(* Logix 5000 project; controller Digital_Interlock_PLC vendor 1 type 14 code 196 rev 37.11; software revision 37.00 *) (continued)
ADD_ON_INSTRUCTION AOI_Sys_Module   (* revision 1.0, vendor Jeremy Medders, ExecutePrescan *)
// Provides detailed module diagnostics and inhibit ability.
VAR_IN_OUT
   Ref_Module : MODULE; {required}   // Name of the module in the I/O tree.
END_VAR
VAR_INPUT
   Inp_Inhibit : BOOL; {access Read Only, visible}   // Command to inhibit the module.
   Inp_Uninhibit : BOOL; {access Read Only, visible}   // Command to uninhibit the module.
END_VAR
VAR_OUTPUT
   Val_EntryStatus : DINT; {access Read Only, visible}   // Specifies the current state of the specified map entry.
   Val_FaultCode : DINT; {access Read Only, visible}   // A number that identifies a module fault, if one occurs.
   Val_FaultInfo : DINT; {access Read Only, visible}   // Provides specific information about the Module object fault code.
   Val_Instance : DINT; {access Read Only, visible}   // Provides the instance number of this module object.
   Val_Mode : DINT; {access Read Only, visible}   // Specifies the current mode of the Module object.
   Sts_Standby : ALIAS FOR Status.0; {access Read Only, visible}   // The controller is powering up.
   Sts_Faulted : ALIAS FOR Status.1; {access Read Only, visible}   // Indicates whether any of the Module object’s connections to the associated module have failed.
   Sts_Validating : ALIAS FOR Status.2; {access Read Only, visible}   // The Module object is verifying Module object integrity prior to establishing connections to the module.
   Sts_Connecting : ALIAS FOR Status.3; {access Read Only, visible}   // The Module object is initiating connections to the module.
   Sts_Connected : ALIAS FOR Status.4; {access Read Only, visible}   // All connections to the module are established and data is transferring.
   Sts_ShuttingDown : ALIAS FOR Status.5; {access Read Only, visible}   // The Module object is in the process of shutting down all connections to the module.
   Sts_Inhibited : ALIAS FOR Status.6; {access Read Only, visible}   // The Module object is inhibited (the inhibit bit in the Mode attribute is set).
   Sts_Waiting : ALIAS FOR Status.7; {access Read Only, visible}   // The parent object upon which this Module object depends is not running.
   Sts_FirmwareUpdating : ALIAS FOR Status.9; {access Read Only, visible}   // Firmware supervisor is attempting to flash the module.
   Sts_Configuring : ALIAS FOR Status.10; {access Read Only, visible}   // Controller is downloading configuration to the module.
   Sts_Disconnected : ALIAS FOR Status.11; {access Read Only, visible}
END_VAR
VAR
   ModeSet : DINT; {access None}
   OSR : BOOL; {access None}
   ESts : DINT; {access None}
   Status : DINT; {access Read Only}
END_VAR

ROUTINE Logic   (* structured text *)
   
   /*
       AO_Sys_Module
       Purpose:
         - Read a module object's status, fault info, and mode
         - One-shot inhibit/uninhibit via Mode bit 2 (0x0004)
         - Decode EntryStatus into HMI-friendly booleans
   */
   
   // --- Snapshot current module diagnostics/state ---
   GSV(Module, Ref_Module, INSTANCE, Val_Instance);
   GSV(Module, Ref_Module, EntryStatus, Val_EntryStatus);
   GSV(Module, Ref_Module, FaultCode, Val_FaultCode);
   GSV(Module, Ref_Module, FaultInfo, Val_FaultInfo);
   GSV(Module, Ref_Module, Mode, Val_Mode);
   
   // --- Rising-edge one-shots for inhibit control (bit 2 of Mode) ---
   // Inhibit: set bit 2
   if (Inp_Inhibit & NOT OSR) then
   	ModeSet := Val_Mode OR 16#0004;
   	SSV(Module, Ref_Module, Mode, ModeSet);
   
   // Uninhibit: clear bit 2
   elsif (Inp_Uninhibit & NOT OSR) then
   	ModeSet := Val_Mode AND 16#FFFB;
   	SSV(Module, Ref_Module, Mode, ModeSet);
   end_if;
   
   // One-shot memory: true for one scan when either command goes high
   OSR := Inp_Inhibit OR Inp_Uninhibit;
   
   /*
   	Entry Status Map
   	• 0x0000: Standby
   	• 0x1000: Faulted
   	• 0x2000: Validating
   	• 0x3000: Connecting
   	• 0x4000: Running
   	• 0x5000: Shutting Down
   	• 0x6000: Inhibited
   	• 0x7000: Waiting
   	• 0x9000: Firmware Updating
   	• 0xA000: Configuring
   */
   ESts := Val_EntryStatus & 16#F000;
   
   // State booleans for HMI/logic
   Sts_Standby := (ESts = 16#0000);
   Sts_Faulted := (ESts = 16#1000);
   Sts_Validating := (ESts = 16#2000);
   Sts_Connecting := (ESts = 16#3000);
   Sts_Connected := (ESts = 16#4000);
   Sts_ShuttingDown := (ESts = 16#5000);
   Sts_Inhibited := (ESts = 16#6000);
   Sts_Waiting := (ESts = 16#7000);
   Sts_FirmwareUpdating := (ESts = 16#9000);
   Sts_Configuring := (ESts = 16#A000);
   Sts_Disconnected := NOT (Sts_Inhibited OR Sts_Connected);
   
END_ROUTINE

ROUTINE Prescan   (* structured text *)
   
   /*
   	AO_Sys_Module
   */
   
   Inp_Inhibit := 0;
   Inp_Uninhibit := 0;
   
   Status := 0;
   
   Val_Instance := 0;
   Val_EntryStatus := 0;
   Val_FaultCode := 0;
   Val_FaultInfo := 0;
   Val_Mode := 0;
   
END_ROUTINE
END_ADD_ON_INSTRUCTION

VAR_GLOBAL   (* controller tags *)
   _DEBUG : BOOL;
   CommsStatus : DINT;
        .3   // LIC comms ok
        .0   // Prefeeder comms ok
        .1   // Stacker comms ok
        .2   // Press comms ok
   CommsStatus_Prefeeder : DINT := 11;
   CommsStatus_Press : DINT;
   CommsStatus_Stacker : DINT;
   EnableLineOptimization : BOOL;
   FaultDetected : BOOL;   // Bool to execute fault routine
   FeedInterruptActive : BOOL;
   FromLIC : UDT_FromLIC;   // Data received from LIC Client
   FromPrefeeder : UDT_EIP_FromPrefeeder;
   FromPress : UDT_EIP_FromPress;
   FromStacker : UDT_EIP_FromStacker;
   HB_ScanCounter : INT := 50;
   HB_Timer1 : TIMER := (PRE := 20);
   HB_Timer2 : TIMER := (PRE := 20);
   HeartBeat : DINT;
   MachineCount : DINT;
   PF_MSG : MESSAGE;
        MessageParameters(ServiceCode := 16#004d, LocalElement := ToPrefeeder.Heartbeat, ...)
   State : UDT_StateContext;
   States : UDT_States;
   ToLIC : UDT_ToLIC;   // Data sent to LIC Client
   ToPrefeeder : UDT_EIP_ToPrefeeder := (Heartbeat := 27);
   ToPress : UDT_EIP_ToPress;
   ToStacker : UDT_EIP_ToStacker := (PrintStation[0].blnSideWaysActive := 1);
END_VAR

PROGRAM Fault_Handler_Program   (* main routine ControllerFaultHandlerRoutine, fault routine CheckSpecificFaultRoutine *)
VAR
   CPU_Scanning : BOOL;   // Identifies when the controller is in prescan.Used t to determine if the fault occurred during prescan or normal scan of the logic
   FaultCode : DINT := 20;
   FaultType : DINT := 4;
   MajorFaultRecord : UDT_FaultRecord;
        .TimeLow   // Stores the fault information in the major_fault_record tag. When you enter a tag that is based on a structure, enter the first member of the tag
   MF_ClearRequestEnable : BOOL;   // allow program to clear this class of fault
   MF_Code : DINT;
   MF_Latched : BOOL;   // Goes true when new fault captured
   MF_Msg : STRING;
   MF_T01_C01 : STR_MajorFault := 'Major Fault T01:C01 - Power-up Fault: Power lost and restored in RUN mode. The controller that is powered on is in Run mode.'; {constant}   // The controller that is powered on is in Run mode.
   MF_T01_C16 : STR_MajorFault := 'Major Fault T01:C16 - Power-up Fault: I/O Communications Configuration fault detected.. I/O communication configuration fault detected.'; {constant}   // I/O communication configuration fault detected.
   MF_T01_C60 : STR_MajorFault := 'Major Fault T01:C60 - Power-up Fault: Non-recoverable fault. The controller detected a nonrecoverable major fault. Diagnostic information can be recovered.'; {constant}   // The controller detected a nonrecoverable major fault. Diagnostic information can be recovered.
   MF_T01_C61 : STR_MajorFault := 'Major Fault T01:C61 - Power-up Fault: Non-recoverable fault with saved diagnostic information. The controller detected a nonrecoverable major fault. Diagnostic information can be recovered.'; {constant}   // The controller detected a nonrecoverable major fault. Diagnostic information can be recovered.
   MF_T03_C16 : STR_MajorFault := 'Major Fault T03:C16 - I/O Fault: I/O module connection failed on required module. A required I/O module connection failed.'; {constant}   // A required I/O module connection failed.
   MF_T03_C23 : STR_MajorFault := 'Major Fault T03:C23 - I/O Fault: At least one required connection not established before going into RUN mode. At least one required connection was not established before going to Run mode.'; {constant}   // At least one required connection was not established before going to Run mode.
   MF_T03_C32 : STR_MajorFault := 'Major Fault T03:C32 - I/O Fault: Controller failed to open an I/O connection to a fault-tolerant I/O module because its partner controller is in a Primary state. The controller failed to open an I/O c'; {constant}   // The controller failed to open an I/O connection to a fault-tolerant I/O module because its partner controller is in a Primary state.
   MF_T03_C94 : STR_MajorFault := 'Minor Fault T03:C94 - I/O Fault: Module RPI overlap detected. The current RPI update of an I/O module overlaps with its previous RPI update.'; {constant}   // The current RPI update of an I/O module overlaps with its previous RPI update.
   MF_Timestamp : DINT;   // UTC seconds/millis, optional timestamp
   MF_Type : DINT;
END_VAR

ROUTINE CheckSpecificFaultRoutine   (* ladder *)
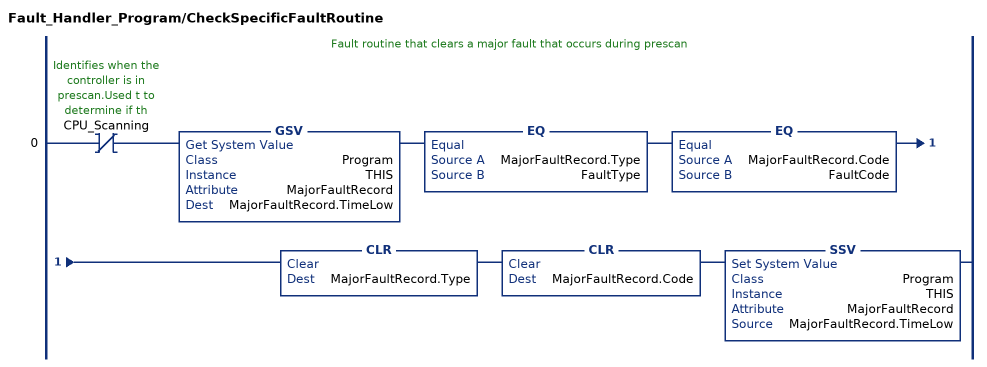
   // Fault routine that clears a major fault that occurs during prescan
   0: XIO(CPU_Scanning)GSV(Program,THIS,MajorFaultRecord,MajorFaultRecord.TimeLow)EQ(MajorFaultRecord.Type,FaultType)EQ(MajorFaultRecord.Code,FaultCode)CLR(MajorFaultRecord.Type)CLR(MajorFaultRecord.Code)SSV(Program,THIS,MajorFaultRecord,MajorFaultRecord.TimeLow);
END_ROUTINE

ROUTINE ControllerFaultHandlerRoutine   (* ladder *)
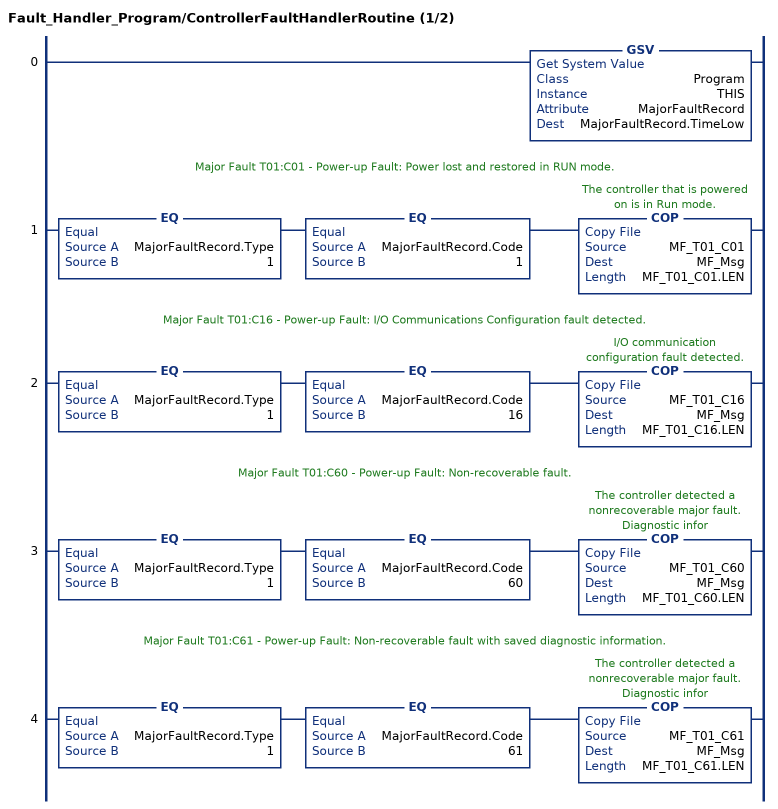
   0: GSV(Program,THIS,MajorFaultRecord,MajorFaultRecord.TimeLow);
   // Major Fault T01:C01 - Power-up Fault: Power lost and restored in RUN mode.
   1: EQ(MajorFaultRecord.Type,1)EQ(MajorFaultRecord.Code,1)COP(MF_T01_C01,MF_Msg,MF_T01_C01.LEN);
   // Major Fault T01:C16 - Power-up Fault: I/O Communications Configuration fault detected.
   2: EQ(MajorFaultRecord.Type,1)EQ(MajorFaultRecord.Code,16)COP(MF_T01_C16,MF_Msg,MF_T01_C16.LEN);
   // Major Fault T01:C60 - Power-up Fault: Non-recoverable fault.
   3: EQ(MajorFaultRecord.Type,1)EQ(MajorFaultRecord.Code,60)COP(MF_T01_C60,MF_Msg,MF_T01_C60.LEN);
   // Major Fault T01:C61 - Power-up Fault: Non-recoverable fault with saved diagnostic information.
   4: EQ(MajorFaultRecord.Type,1)EQ(MajorFaultRecord.Code,61)COP(MF_T01_C61,MF_Msg,MF_T01_C61.LEN);
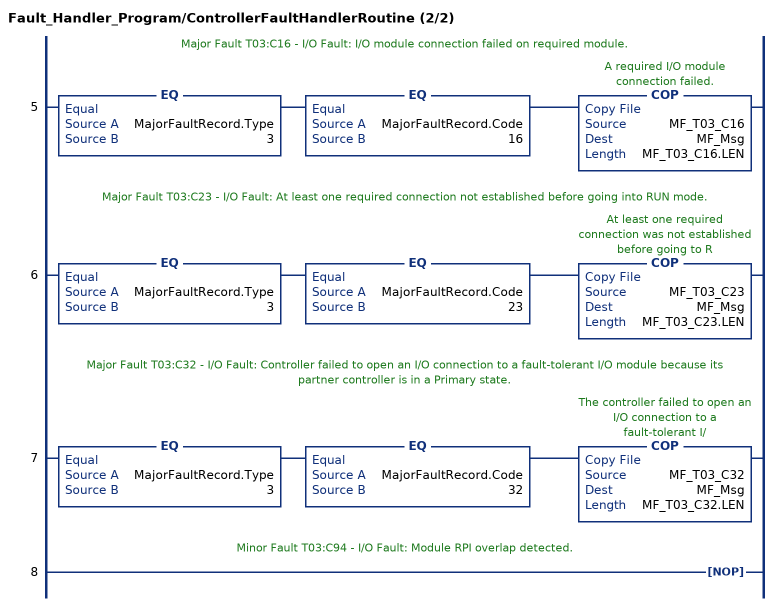
   // Major Fault T03:C16 - I/O Fault: I/O module connection failed on required module.
   5: EQ(MajorFaultRecord.Type,3)EQ(MajorFaultRecord.Code,16)COP(MF_T03_C16,MF_Msg,MF_T03_C16.LEN);
   // Major Fault T03:C23 - I/O Fault: At least one required connection not established before going into RUN mode.
   6: EQ(MajorFaultRecord.Type,3)EQ(MajorFaultRecord.Code,23)COP(MF_T03_C23,MF_Msg,MF_T03_C23.LEN);
   // Major Fault T03:C32 - I/O Fault: Controller failed to open an I/O connection to a fault-tolerant I/O module because its partner controller is in a Primary state.
   7: EQ(MajorFaultRecord.Type,3)EQ(MajorFaultRecord.Code,32)COP(MF_T03_C32,MF_Msg,MF_T03_C32.LEN);
   // Minor Fault T03:C94 - I/O Fault: Module RPI overlap detected.
   8: NOP();
END_ROUTINE
END_PROGRAM

PROGRAM MainProgram   (* main routine MainRoutine *)
VAR
   AlwaysTrue : BOOL := 1; {constant}
   AnyFault : BOOL;
   BR1_Health : UDT_DeviceHealth;
   BR2_Health : UDT_DeviceHealth;
   CmdEdge_Interrupt : BOOL;
   CmdEdge_Reconfig : BOOL;
   CmdEdge_Reset : BOOL;
   CmdEdge_Start : BOOL;
   CmdEdge_Stop : BOOL;
   CmdId_Desired : DINT;
   CmdId_Last : DINT;
   CN1_Health : UDT_DeviceHealth;
   CN2_Health : UDT_DeviceHealth;
   CommandEnum : UDT_CommandEnum;
   CommsHealthy : BOOL;   // Heartbeat Ok between peer machines
   DesiredCommand : DINT;   // From LIC Client
   EndCriteriaMet : BOOL;
   GuardsOk : BOOL;
   HeartBeatB : BOOL := 1;
   HoldClear : BOOL;
   HWReady : BOOL;   // Machines present and communicating
   MajorFaultRec : UDT_FaultRecord;
   ONS_CmdId : BOOL;
   PermissivesOk : BOOL;   // (safety, e-stops, power, guards
   PF1_Health : UDT_DeviceHealth := (DeviceConfigured := 1);
   PF2_Health : UDT_DeviceHealth;
   PL1_Health : UDT_DeviceHealth;
   PL2_Health : UDT_DeviceHealth;
   PowerOk : BOOL;
   PR1_Health : UDT_DeviceHealth;
   PR2_Health : UDT_DeviceHealth;
   SafetyChain_OK : BOOL;
   SR1_Health : UDT_DeviceHealth;
   SR2_Health : UDT_DeviceHealth;
   ST1_Health : UDT_DeviceHealth := (DeviceConfigured := 1);
   ST2_Health : UDT_DeviceHealth;
   TaskPeriod_ms : DINT := 10; {constant}   // must match periodic task ms
   TB1_Health : UDT_DeviceHealth;
   TB2_Health : UDT_DeviceHealth;
   Tmr_Hold : TIMER := (PRE := 10000);
   Tmr_Init : TIMER := (PRE := 3000);
   Tmr_Running : TIMER := (PRE := 5000);
END_VAR

ROUTINE DataRoutingRoutine   (* structured text *)
   
   /******************** 	DATA MAPPING	********************/
   
   ST1:O.Data[0] := ToStacker.Heartbeat;										// Press -> Stacker
   ST1:O.Data[1] := ToStacker.CommandedSpeed;									// Press -> Stacker
   ST1:O.Data[2] := ToStacker.PressCurrentSpeed;								// Press -> Stacker
   ST1:O.Data[3].0 := ToStacker.RollInPermissive;								// Press -> Stacker
   ST1:O.Data[3].1 := ToStacker.RunPermissive;									// Press -> Stacker
   ST1:O.Data[3].2 := ToStacker.VOSReset;										// Press -> Stacker
   ST1:O.Data[3].3 := ToStacker.VOSStart;										// Press -> Stacker
   ST1:O.Data[3].4 := ToStacker.SheetCountPulseStatus;							// Press -> Stacker
   ST1:O.Data[3].5 := ToStacker.DieCutter.blnRegistrationActive;				// Press -> Stacker
   ST1:O.Data[3].6 := ToStacker.DieCutter.blnSidewaysAcitve;					// Press -> Stacker
   ST1:O.Data[3].7 := ToStacker.DieCutter.blnSpeedChangeActive;				// Press -> Stacker
   ST1:O.Data[3].8 := ToStacker.PrintStation[0].blnRegistrationActive;			// Press -> Stacker
   ST1:O.Data[3].9 := ToStacker.PrintStation[1].blnRegistrationActive;			// Press -> Stacker
   ST1:O.Data[3].10 := ToStacker.PrintStation[2].blnRegistrationActive;		// Press -> Stacker
   ST1:O.Data[3].11 := ToStacker.PrintStation[3].blnRegistrationActive;		// Press -> Stacker
   ST1:O.Data[3].12 := ToStacker.PrintStation[4].blnRegistrationActive;		// Press -> Stacker
   ST1:O.Data[3].13 := ToStacker.PrintStation[5].blnRegistrationActive;		// Press -> Stacker
   ST1:O.Data[3].14 := ToStacker.PrintStation[6].blnRegistrationActive;		// Press -> Stacker
   ST1:O.Data[3].15 := ToStacker.PrintStation[0].blnSideWaysActive;			// Press -> Stacker
   ST1:O.Data[3].16 := ToStacker.PrintStation[1].blnSideWaysActive;			// Press -> Stacker
   ST1:O.Data[3].17 := ToStacker.PrintStation[2].blnSideWaysActive;			// Press -> Stacker
   ST1:O.Data[3].18 := ToStacker.PrintStation[3].blnSideWaysActive;			// Press -> Stacker
   ST1:O.Data[3].19 := ToStacker.PrintStation[4].blnSideWaysActive;			// Press -> Stacker
   ST1:O.Data[3].20 := ToStacker.PrintStation[5].blnSideWaysActive;			// Press -> Stacker
   ST1:O.Data[3].21 := ToStacker.PrintStation[6].blnSideWaysActive;			// Press -> Stacker
   ST1:O.Data[3].22 := ToStacker.DownstreamReady;								// LIC -> Stacker
   ST1:O.Data[4] := ToStacker.DieCutter.uiActualSpeedKpm;						// Press -> Stacker
   ST1:O.Data[5] := ToStacker.DieCutter.fltActualRegisterPosition;				// Press -> Stacker
   ST1:O.Data[6] := ToStacker.DieCutter.fltActualSidewaysPosition;				// Press -> Stacker
   ST1:O.Data[7] := ToStacker.PrintStation[0].fltActualRegisterPosition;		// Press -> Stacker
   ST1:O.Data[8] := ToStacker.PrintStation[1].fltActualRegisterPosition;		// Press -> Stacker
   ST1:O.Data[9] := ToStacker.PrintStation[2].fltActualRegisterPosition;		// Press -> Stacker
   ST1:O.Data[10] := ToStacker.PrintStation[3].fltActualRegisterPosition;		// Press -> Stacker
   ST1:O.Data[11] := ToStacker.PrintStation[4].fltActualRegisterPosition;		// Press -> Stacker
   ST1:O.Data[12] := ToStacker.PrintStation[5].fltActualRegisterPosition;		// Press -> Stacker
   ST1:O.Data[13] := ToStacker.PrintStation[6].fltActualRegisterPosition;		// Press -> Stacker
   ST1:O.Data[14] := ToStacker.PrintStation[0].fltActualSidewaysPosition;		// Press -> Stacker
   ST1:O.Data[15] := ToStacker.PrintStation[1].fltActualSidewaysPosition;		// Press -> Stacker
   ST1:O.Data[16] := ToStacker.PrintStation[2].fltActualSidewaysPosition;		// Press -> Stacker
   ST1:O.Data[17] := ToStacker.PrintStation[3].fltActualSidewaysPosition;		// Press -> Stacker
   ST1:O.Data[18] := ToStacker.PrintStation[4].fltActualSidewaysPosition;		// Press -> Stacker
   ST1:O.Data[19] := ToStacker.PrintStation[5].fltActualSidewaysPosition;		// Press -> Stacker
   ST1:O.Data[20] := ToStacker.PrintStation[6].fltActualSidewaysPosition;		// Press -> Stacker
   ST1:O.Data[20] := ToStacker.CommsStatus;									// Interlock -> Stacker
   /*-------------------------------------------------------------*/
   
   FromStacker.Heartbeat := ST1:I.Data[6];										// Stacker -> Press
   FromStacker.CurrentSpeed := ST1:I.Data[7];									// Stacker -> Press
   FromStacker.PatternMaxSpeed := ST1:I.Data[8];								// Stacker -> Press
   FromStacker.FillPercentage := ST1:I.Data[9];								// Stacker -> Press
   FromStacker.RunPermissive := ST1:I.Data[10].0;								// Stacker -> Press
   FromStacker.FeedRestart := ST1:I.Data[10].1; 								// Stacker -> Press
   FromStacker.RolledOutStatus := ST1:I.Data[10].2; 							// Stacker -> Press
   FromStacker.FeedInterruptStatus := ST1:I.Data[10].3;						// Stacker -> Press
   FromStacker.DieCutter.blnFast := ST1:I.Data[10].4;							// Stacker -> Press
   FromStacker.DieCutter.blnSlow := ST1:I.Data[10].5;							// Stacker -> Press
   FromStacker.DieCutter.blnRegisterAdjustRq := ST1:I.Data[10].6;				// Stacker -> Press
   FromStacker.DieCutter.blnRegisterStopAdjustRq := ST1:I.Data[10].7;			// Stacker -> Press
   FromStacker.DieCutter.blnSidewaysAdjustRq := ST1:I.Data[10].8;				// Stacker -> Press
   FromStacker.DieCutter.blnSidewaysStopAdjustRq := ST1:I.Data[10].9;			// Stacker -> Press
   FromStacker.DieCutter.blnSpeedChangeRq := ST1:I.Data[10].10;				// Stacker -> Press
   FromStacker.DieCutter.blnSpeedChangeStopRq := ST1:I.Data[10].11;			// Stacker -> Press
   FromStacker.PrintStation[0].blnRegisterAdjustRq := ST1:I.Data[10].12;		// Stacker -> Press
   FromStacker.PrintStation[1].blnRegisterAdjustRq := ST1:I.Data[10].13;		// Stacker -> Press
   FromStacker.PrintStation[2].blnRegisterAdjustRq := ST1:I.Data[10].14;		// Stacker -> Press
   FromStacker.PrintStation[3].blnRegisterAdjustRq := ST1:I.Data[10].15;		// Stacker -> Press
   FromStacker.PrintStation[4].blnRegisterAdjustRq := ST1:I.Data[10].16;		// Stacker -> Press
   FromStacker.PrintStation[5].blnRegisterAdjustRq := ST1:I.Data[10].17;		// Stacker -> Press
   FromStacker.PrintStation[6].blnRegisterAdjustRq := ST1:I.Data[10].18;		// Stacker -> Press
   FromStacker.PrintStation[0].blnSidewaysAdjustRq := ST1:I.Data[10].19;		// Stacker -> Press
   FromStacker.PrintStation[1].blnSidewaysAdjustRq := ST1:I.Data[10].20;		// Stacker -> Press
   FromStacker.PrintStation[2].blnSidewaysAdjustRq := ST1:I.Data[10].21;		// Stacker -> Press
   FromStacker.PrintStation[3].blnSidewaysAdjustRq := ST1:I.Data[10].22;		// Stacker -> Press
   FromStacker.PrintStation[4].blnSidewaysAdjustRq := ST1:I.Data[10].23;		// Stacker -> Press
   FromStacker.PrintStation[5].blnSidewaysAdjustRq := ST1:I.Data[10].24;		// Stacker -> Press
   FromStacker.PrintStation[6].blnSidewaysAdjustRq := ST1:I.Data[10].25;		// Stacker -> Press
   FromStacker.PrintStation[0].blnRegisterStopAdjustRq := ST1:I.Data[10].26;	// Stacker -> Press
   FromStacker.PrintStation[1].blnRegisterStopAdjustRq := ST1:I.Data[10].27;	// Stacker -> Press
   FromStacker.PrintStation[2].blnRegisterStopAdjustRq := ST1:I.Data[10].28;	// Stacker -> Press
   FromStacker.PrintStation[3].blnRegisterStopAdjustRq := ST1:I.Data[10].29;	// Stacker -> Press
   FromStacker.PrintStation[4].blnRegisterStopAdjustRq := ST1:I.Data[10].30;	// Stacker -> Press
   FromStacker.PrintStation[5].blnRegisterStopAdjustRq := ST1:I.Data[10].31;	// Stacker -> Press
   FromStacker.PrintStation[6].blnRegisterStopAdjustRq := ST1:I.Data[11].0;	// Stacker -> Press
   FromStacker.PrintStation[0].blnSidewaysStopAdjustRq := ST1:I.Data[11].1;	// Stacker -> Press
   FromStacker.PrintStation[1].blnSidewaysStopAdjustRq := ST1:I.Data[11].2;	// Stacker -> Press
   FromStacker.PrintStation[2].blnSidewaysStopAdjustRq := ST1:I.Data[11].3;	// Stacker -> Press
   FromStacker.PrintStation[3].blnSidewaysStopAdjustRq := ST1:I.Data[11].4;	// Stacker -> Press
   FromStacker.PrintStation[4].blnSidewaysStopAdjustRq := ST1:I.Data[11].5;	// Stacker -> Press
   FromStacker.PrintStation[5].blnSidewaysStopAdjustRq := ST1:I.Data[11].6;	// Stacker -> Press
   FromStacker.PrintStation[6].blnSidewaysStopAdjustRq := ST1:I.Data[11].7;	// Stacker -> Press
   FromStacker.DieCutter.uiDesiredSpeedKpm := ST1:I.Data[12];					// Stacker -> Press
   FromStacker.DieCutter.fltDesiredRegisterAdjust := ST1:I.Data[13];			// Stacker -> Press
   FromStacker.PrintStation[0].fltDesiredRegisterAdjust := ST1:I.Data[14];		// Stacker -> Press
   FromStacker.PrintStation[1].fltDesiredRegisterAdjust := ST1:I.Data[15];		// Stacker -> Press
   FromStacker.PrintStation[2].fltDesiredRegisterAdjust := ST1:I.Data[16];		// Stacker -> Press
   FromStacker.PrintStation[3].fltDesiredRegisterAdjust := ST1:I.Data[17];		// Stacker -> Press
   FromStacker.PrintStation[4].fltDesiredRegisterAdjust := ST1:I.Data[18];		// Stacker -> Press
   FromStacker.PrintStation[5].fltDesiredRegisterAdjust := ST1:I.Data[19];		// Stacker -> Press
   FromStacker.PrintStation[6].fltDesiredRegisterAdjust := ST1:I.Data[20];		// Stacker -> Press
   FromStacker.DieCutter.fltDesiredSidewaysAdjust := ST1:I.Data[21];			// Stacker -> Press
   FromStacker.PrintStation[0].fltDesiredSidewaysAdjust := ST1:I.Data[22];		// Stacker -> Press
   FromStacker.PrintStation[1].fltDesiredSidewaysAdjust := ST1:I.Data[23];		// Stacker -> Press
   FromStacker.PrintStation[2].fltDesiredSidewaysAdjust := ST1:I.Data[24];		// Stacker -> Press
   FromStacker.PrintStation[3].fltDesiredSidewaysAdjust := ST1:I.Data[25];		// Stacker -> Press
   FromStacker.PrintStation[4].fltDesiredSidewaysAdjust := ST1:I.Data[26];		// Stacker -> Press
   FromStacker.PrintStation[5].fltDesiredSidewaysAdjust := ST1:I.Data[27];		// Stacker -> Press
   FromStacker.PrintStation[6].fltDesiredSidewaysAdjust := ST1:I.Data[28];		// Stacker -> Press
   FromStacker.Spare1 := ST1:I.Data[29];
   FromStacker.Spare2 :=  ST1:I.Data[30];
   /*-------------------------------------------------------------*/
   
   PR1:O.Data[0].0 := ToPress.AuxTamperAirRight;			// Pre-Feeder -> Press
   PR1:O.Data[0].1 := ToPress.AuxTamperAirLeft;			// Pre-Feeder -> Press
   PR1:O.Data[0].2 := ToPress.BackstopInhibit;				// Pre-Feeder -> Press
   PR1:O.Data[0].3 := ToPress.CallForStack;				// Pre-Feeder -> Press
   PR1:O.Data[0].4 := ToPress.ExtendoUpDown;				// Pre-Feeder -> Press
   PR1:O.Data[0].5 := ToPress.EstopFeedbackChannel1;		// Pre-Feeder -> Press
   PR1:O.Data[0].6 := ToPress.EstopFeedbackChannel2;		// Pre-Feeder -> Press
   PR1:O.Data[0].7 := ToPress.FeedBoardOk;					// Pre-Feeder -> Press
   PR1:O.Data[0].8 := ToPress.MachineOpenCloseDisable;		// Pre-Feeder -> Press
   PR1:O.Data[0].9 := ToPress.OpenMachineOk;				// Pre-Feeder -> Press
   PR1:O.Data[0].10 := ToPress.ReadyForSetup;				// Pre-Feeder -> Press
   PR1:O.Data[0].11 := ToPress.ReadyToRaise;				// Pre-Feeder -> Press
   PR1:O.Data[0].12 := ToPress.RunEmpty;					// Pre-Feeder -> Press
   PR1:O.Data[0].13 := ToPress.RunForward;					// Pre-Feeder -> Press
   PR1:O.Data[0].14 := ToPress.RunReverse;					// Pre-Feeder -> Press
   PR1:O.Data[0].15 := ToPress.TamperInterrupt;			// Pre-Feeder -> Press
   PR1:O.Data[0].16 := ToPress.Empty;						// Pre-Feeder -> Press
   PR1:O.Data[0].17 := ToPress.FeedInterrupt;				// Pre-Feeder -> Press
   PR1:O.Data[0].18 := ToPress.Spare;						// Pre-Feeder -> Press
   PR1:O.Data[1] := ToPress.CurrentSpeed;					// Pre-Feeder -> Press
   PR1:O.Data[2] := ToPress.PatternMaxSpeed;				// Pre-Feeder -> Press
   PR1:O.Data[3] := ToPress.Heartbeat_Echo_Prefeeder;		// Pre-Feeder -> Press
   PR1:O.Data[4] := ToPress.Spare1;						// Pre-Feeder -> Press
   PR1:O.Data[5] := ToPress.Spare2;						// Pre-Feeder -> Press
   PR1:O.Data[6] := ToPress.Heartbeat_Echo_Stacker;		// Stacker -> Press
   PR1:O.Data[7] := ToPress.CurrentSpeed;					// Stacker -> Press
END_ROUTINE

ROUTINE HeartbeatRoutine   (* ladder *)
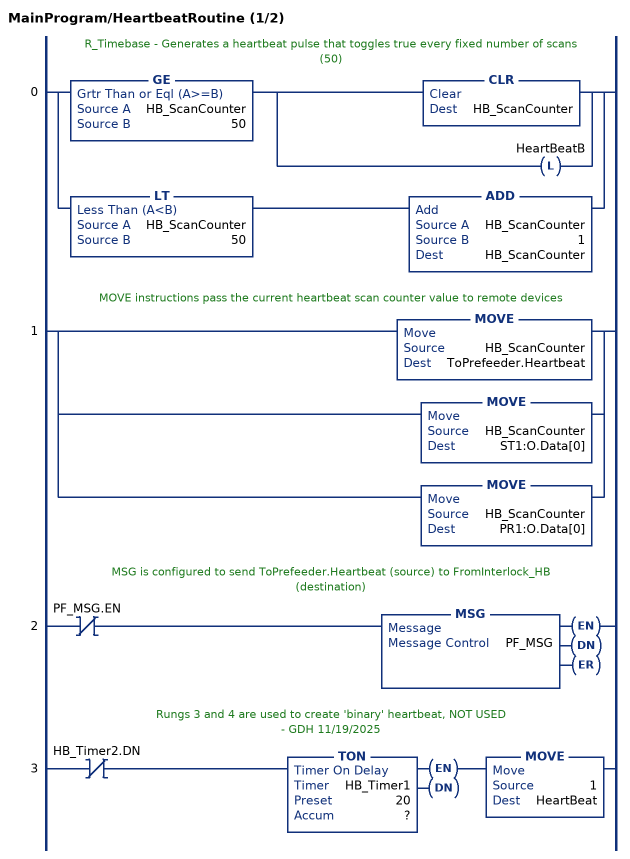
   // R_Timebase - Generates a heartbeat pulse that toggles true every fixed number of scans (50)
   0: [GE(HB_ScanCounter,50) [CLR(HB_ScanCounter) ,OTL(HeartBeatB) ] ,LT(HB_ScanCounter,50) ADD(HB_ScanCounter,1,HB_ScanCounter) ];
   // MOVE instructions pass the current heartbeat scan counter value to remote devices
   1: [MOVE(HB_ScanCounter,ToPrefeeder.Heartbeat) ,MOVE(HB_ScanCounter,ST1:O.Data[0]) ,MOVE(HB_ScanCounter,PR1:O.Data[0]) ];
   // MSG is configured to send ToPrefeeder.Heartbeat (source) to FromInterlock_HB (destination)
   2: XIO(PF_MSG.EN)MSG(PF_MSG);
   // Rungs 3 and 4 are used to create 'binary' heartbeat, NOT USED
   // - GDH 11/19/2025
   3: XIO(HB_Timer2.DN)TON(HB_Timer1,?,?)MOVE(1,HeartBeat);
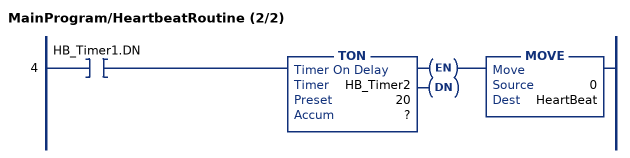
   4: XIC(HB_Timer1.DN)TON(HB_Timer2,?,?)MOVE(0,HeartBeat);
END_ROUTINE

ROUTINE MainRoutine   (* ladder *)
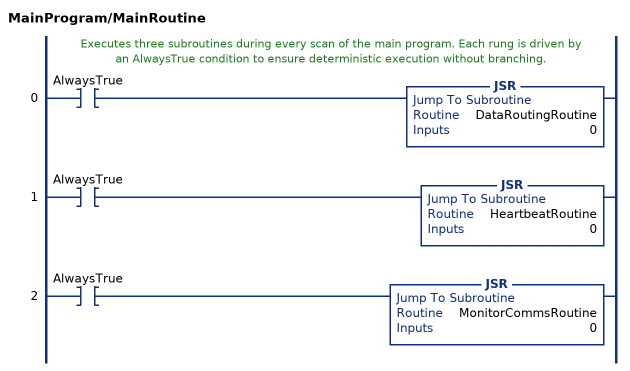
   // Executes three subroutines during every scan of the main program. Each rung is driven by an AlwaysTrue condition to ensure deterministic execution without branching.
   0: XIC(AlwaysTrue)JSR(DataRoutingRoutine,0);
   1: XIC(AlwaysTrue)JSR(HeartbeatRoutine,0);
   2: XIC(AlwaysTrue)JSR(MonitorCommsRoutine,0);
END_ROUTINE

ROUTINE MonitorCommsRoutine   (* structured text *)
   // -------------Press--------------------//
   if PR1_Health.DeviceConfigured then
   	GSV(Module,PR1,EntryStatus,PR1_Health.EntryStatus);
   	GSV(Module,PR1,FaultCode,PR1_Health.FaultCode);
   	GSV(Module,PR1,FaultInfo,PR1_Health.FaultInfo);
   end_if;
   
   // -------------Prefeeder-----------------//
   if PF1_Health.DeviceConfigured then
   	GSV(Module,PF1,EntryStatus,PF1_Health.EntryStatus);
   	GSV(Module,PF1,FaultCode,PF1_Health.FaultCode);
   	GSV(Module,PF1,FaultInfo,PF1_Health.FaultInfo);
   end_if;
   
   if ST1_Health.DeviceConfigured then
   	GSV(Module,ST1,EntryStatus,ST1_Health.EntryStatus);
   	GSV(Module,ST1,FaultCode,ST1_Health.FaultCode);
   	GSV(Module,ST1,FaultInfo,ST1_Health.FaultInfo);
   end_if;
   
   
   //if PF2_Health.DeviceConfigured then
   //	GSV(Module,PF2,EntryStatus,PF2_Health.EntryStatus);
   //	GSV(Module,PF2,FaultCode,PF2_Health.FaultCode);
   //	GSV(Module,PF2,FaultInfo,PF2_Health.FaultInfo);
   //end_if;
   
   // -------------Stacker-----------------//
   //if ST2_Health.DeviceConfigured then
   //	GSV(Module,ST2,EntryStatus,ST2_Health.EntryStatus);
   //	GSV(Module,ST2,FaultCode,ST2_Health.FaultCode);
   //	GSV(Module,ST2,FaultInfo,ST2_Health.FaultInfo);
   //end_if;
   
   
   //// -------------Conveyor-----------------//
   //if CN1_Health.DeviceConfigured then
   //	GSV(Module,CN1,EntryStatus,CN1_Health.EntryStatus);
   //	GSV(Module,CN1,FaultCode,CN1_Health.FaultCode);
   //	GSV(Module,CN1,FaultInfo,CN1_Health.FaultInfo);
   //end_if;
   
   //if CN2_Health.DeviceConfigured then
   //	GSV(Module,CN2,EntryStatus,CN2_Health.EntryStatus);
   //	GSV(Module,CN2,FaultCode,CN2_Health.FaultCode);
   //	GSV(Module,CN2,FaultInfo,CN2_Health.FaultInfo);
   //end_if;
   
   
   
   //if PR2_Health.DeviceConfigured then
   //	GSV(Module,PR2,EntryStatus,PR2_Health.EntryStatus);
   //	GSV(Module,PR2,FaultCode,PR2_Health.FaultCode);
   //	GSV(Module,PR2,FaultInfo,PR2_Health.FaultInfo);
   //end_if;
   
   //// -------------Strapper-----------------//
   //if SR1_Health.DeviceConfigured then
   //	GSV(Module,SR1,EntryStatus,SR1_Health.EntryStatus);
   //	GSV(Module,SR1,FaultCode,SR1_Health.FaultCode);
   //	GSV(Module,SR1,FaultInfo,SR1_Health.FaultInfo);
   //end_if;
   
   //if SR2_Health.DeviceConfigured then
   //	GSV(Module,SR2,EntryStatus,SR2_Health.EntryStatus);
   //	GSV(Module,SR2,FaultCode,SR2_Health.FaultCode);
   //	GSV(Module,SR2,FaultInfo,SR2_Health.FaultInfo);
   //end_if;
   
   //// -------------Twin Bow Slitter--------//
   //if TB1_Health.DeviceConfigured then
   //	GSV(Module,TB1,EntryStatus,TB1_Health.EntryStatus);
   //	GSV(Module,TB1,FaultCode,TB1_Health.FaultCode);
   //	GSV(Module,TB1,FaultInfo,TB1_Health.FaultInfo);
   //end_if;
   
   //if TB2_Health.DeviceConfigured then
   //	GSV(Module,TB2,EntryStatus,TB2_Health.EntryStatus);
   //	GSV(Module,TB2,FaultCode,TB2_Health.FaultCode);
   //	GSV(Module,TB2,FaultInfo,TB2_Health.FaultInfo);
   //end_if;
   
   //// -------------Breaker-----------------//
   //if BR1_Health.DeviceConfigured then
   //	GSV(Module,BR1,EntryStatus,BR1_Health.EntryStatus);
   //	GSV(Module,BR1,FaultCode,BR1_Health.FaultCode);
   //	GSV(Module,BR1,FaultInfo,BR1_Health.FaultInfo);
   //end_if;
   
   //if BR2_Health.DeviceConfigured then
   //	GSV(Module,BR2,EntryStatus,BR2_Health.EntryStatus);
   //	GSV(Module,BR2,FaultCode,BR2_Health.FaultCode);
   //	GSV(Module,BR2,FaultInfo,BR2_Health.FaultInfo);
   //end_if;
   
   //// -------------Palletizer--------------//
   //if PL1_Health.DeviceConfigured then
   //	GSV(Module,PL1,EntryStatus,PL1_Health.EntryStatus);
   //	GSV(Module,PL1,FaultCode,PL1_Health.FaultCode);
   //	GSV(Module,PL1,FaultInfo,PL1_Health.FaultInfo);
   //end_if;
   
   //if PL2_Health.DeviceConfigured then
   //	GSV(Module,PL2,EntryStatus,PL2_Health.EntryStatus);
   //	GSV(Module,PL2,FaultCode,PL2_Health.FaultCode);
   //	GSV(Module,PL2,FaultInfo,PL2_Health.FaultInfo);
   //end_if;
END_ROUTINE
END_PROGRAM
